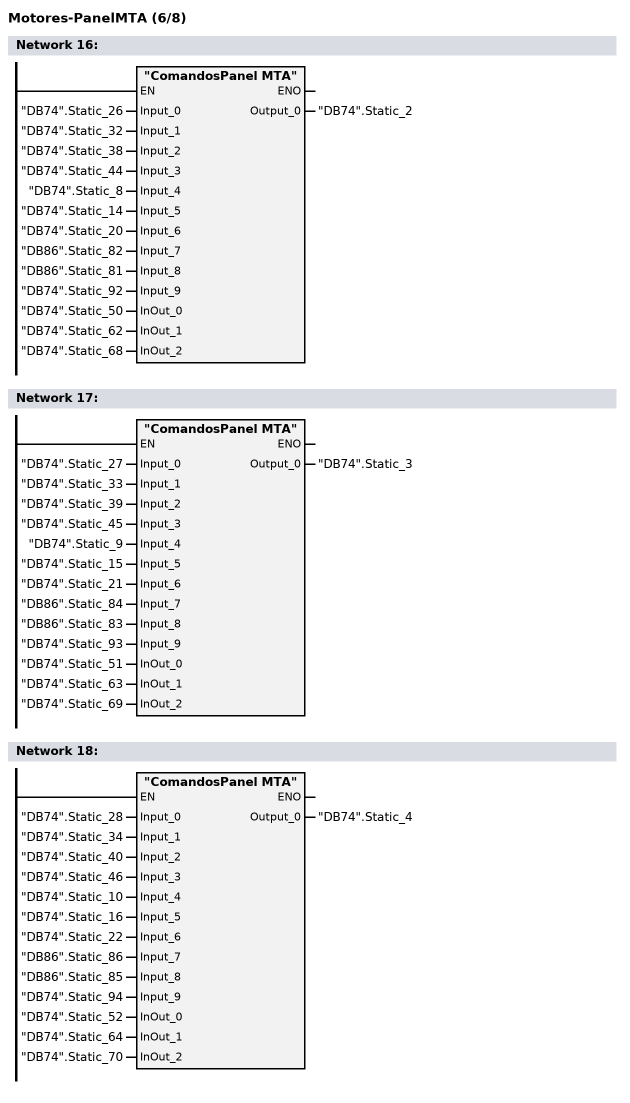
   RUNG wire#powerrail
      "ComandosPanel MTA"(Input_0 := "DB74".Static_26, Input_1 := "DB74".Static_32, Input_2 := "DB74".Static_38, Input_3 := "DB74".Static_44, Input_4 := "DB74".Static_8, Input_5 := "DB74".Static_14, Input_6 := "DB74".Static_20, Input_7 := "DB86".Static_82, Input_8 := "DB86".Static_81, Input_9 := "DB74".Static_92, Output_0 => "DB74".Static_2, InOut_0 := "DB74".Static_50, InOut_1 := "DB74".Static_62, InOut_2 := "DB74".Static_68)
   END_RUNG
   // the same network as SCL:
   "ComandosPanel MTA"(Input_0 := "DB74".Static_26,
                       Input_1 := "DB74".Static_32,
                       Input_2 := "DB74".Static_38,
                       Input_3 := "DB74".Static_44,
                       Input_4 := "DB74".Static_8,
                       Input_5 := "DB74".Static_14,
                       Input_6 := "DB74".Static_20,
                       Input_7 := "DB86".Static_82,
                       Input_8 := "DB86".Static_81,
                       Input_9 := "DB74".Static_92,
                       InOut_0 := "DB74".Static_50,
                       InOut_1 := "DB74".Static_62,
                       InOut_2 := "DB74".Static_68,
                       Output_0 => "DB74".Static_2);
END_REGION

REGION Network 17
   RUNG wire#powerrail
      "ComandosPanel MTA"(Input_0 := "DB74".Static_27, Input_1 := "DB74".Static_33, Input_2 := "DB74".Static_39, Input_3 := "DB74".Static_45, Input_4 := "DB74".Static_9, Input_5 := "DB74".Static_15, Input_6 := "DB74".Static_21, Input_7 := "DB86".Static_84, Input_8 := "DB86".Static_83, Input_9 := "DB74".Static_93, Output_0 => "DB74".Static_3, InOut_0 := "DB74".Static_51, InOut_1 := "DB74".Static_63, InOut_2 := "DB74".Static_69)
   END_RUNG
   // the same network as SCL:
   "ComandosPanel MTA"(Input_0 := "DB74".Static_27,
                       Input_1 := "DB74".Static_33,
                       Input_2 := "DB74".Static_39,
                       Input_3 := "DB74".Static_45,
                       Input_4 := "DB74".Static_9,
                       Input_5 := "DB74".Static_15,
                       Input_6 := "DB74".Static_21,
                       Input_7 := "DB86".Static_84,
                       Input_8 := "DB86".Static_83,
                       Input_9 := "DB74".Static_93,
                       InOut_0 := "DB74".Static_51,
                       InOut_1 := "DB74".Static_63,
                       InOut_2 := "DB74".Static_69,
                       Output_0 => "DB74".Static_3);
END_REGION

REGION Network 18
   RUNG wire#powerrail
      "ComandosPanel MTA"(Input_0 := "DB74".Static_28, Input_1 := "DB74".Static_34, Input_2 := "DB74".Static_40, Input_3 := "DB74".Static_46, Input_4 := "DB74".Static_10, Input_5 := "DB74".Static_16, Input_6 := "DB74".Static_22, Input_7 := "DB86".Static_86, Input_8 := "DB86".Static_85, Input_9 := "DB74".Static_94, Output_0 => "DB74".Static_4, InOut_0 := "DB74".Static_52, InOut_1 := "DB74".Static_64, InOut_2 := "DB74".Static_70)
   END_RUNG
   // the same network as SCL:
   "ComandosPanel MTA"(Input_0 := "DB74".Static_28,
                       Input_1 := "DB74".Static_34,
                       Input_2 := "DB74".Static_40,
                       Input_3 := "DB74".Static_46,
                       Input_4 := "DB74".Static_10,
                       Input_5 := "DB74".Static_16,
                       Input_6 := "DB74".Static_22,
                       Input_7 := "DB86".Static_86,
                       Input_8 := "DB86".Static_85,
                       Input_9 := "DB74".Static_94,
                       InOut_0 := "DB74".Static_52,
                       InOut_1 := "DB74".Static_64,
                       InOut_2 := "DB74".Static_70,
                       Output_0 => "DB74".Static_4);
END_REGION

REGION Network 19
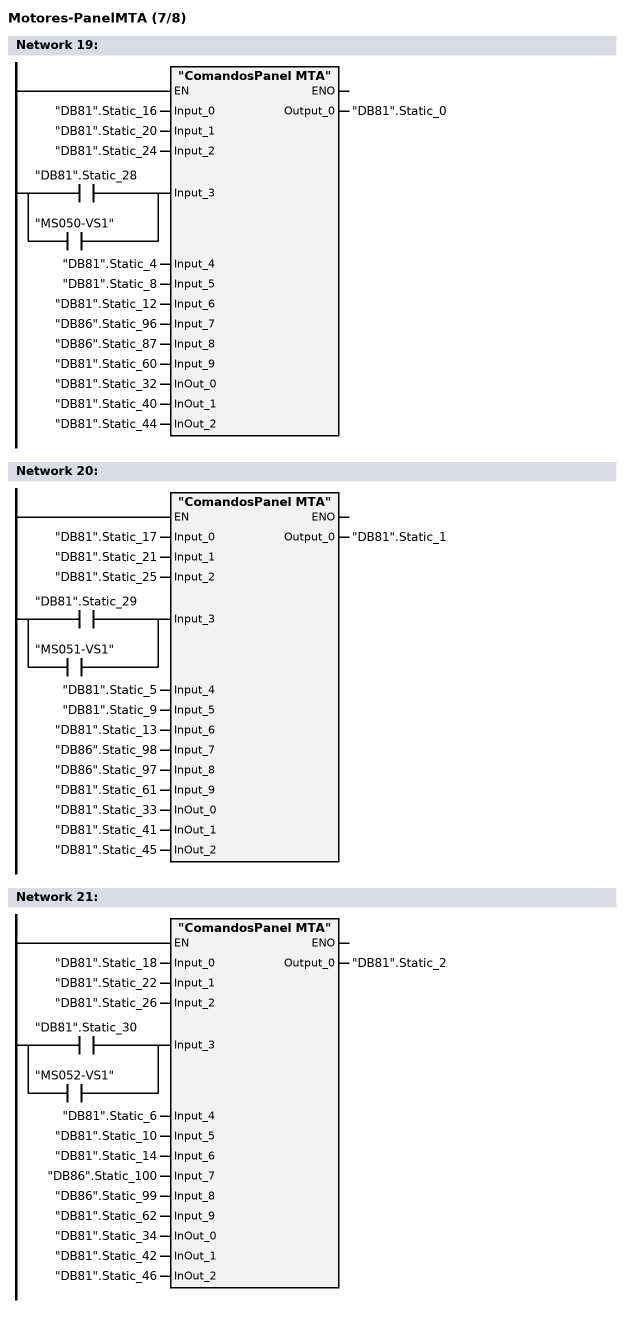
   RUNG wire#powerrail
      "ComandosPanel MTA"(Input_0 := "DB81".Static_16, Input_1 := "DB81".Static_20, Input_2 := "DB81".Static_24, Input_3 := wire#w1, Input_4 := "DB81".Static_4, Input_5 := "DB81".Static_8, Input_6 := "DB81".Static_12, Input_7 := "DB86".Static_96, Input_8 := "DB86".Static_87, Input_9 := "DB81".Static_60, Output_0 => "DB81".Static_0, InOut_0 := "DB81".Static_32, InOut_1 := "DB81".Static_40, InOut_2 := "DB81".Static_44)
   END_RUNG
   RUNG wire#powerrail
      Contact( "DB81".Static_28 )
   END_RUNG wire#w1
   RUNG wire#powerrail
      Contact( "MS050-VS1" )
   END_RUNG wire#w1
   // the same network as SCL:
   "ComandosPanel MTA"(Input_0 := "DB81".Static_16,
                       Input_1 := "DB81".Static_20,
                       Input_2 := "DB81".Static_24,
                       Input_3 := "DB81".Static_28 OR "MS050-VS1",
                       Input_4 := "DB81".Static_4,
                       Input_5 := "DB81".Static_8,
                       Input_6 := "DB81".Static_12,
                       Input_7 := "DB86".Static_96,
                       Input_8 := "DB86".Static_87,
                       Input_9 := "DB81".Static_60,
                       InOut_0 := "DB81".Static_32,
                       InOut_1 := "DB81".Static_40,
                       InOut_2 := "DB81".Static_44,
                       Output_0 => "DB81".Static_0);
END_REGION

REGION Network 20
   RUNG wire#powerrail
      "ComandosPanel MTA"(Input_0 := "DB81".Static_17, Input_1 := "DB81".Static_21, Input_2 := "DB81".Static_25, Input_3 := wire#w1, Input_4 := "DB81".Static_5, Input_5 := "DB81".Static_9, Input_6 := "DB81".Static_13, Input_7 := "DB86".Static_98, Input_8 := "DB86".Static_97, Input_9 := "DB81".Static_61, Output_0 => "DB81".Static_1, InOut_0 := "DB81".Static_33, InOut_1 := "DB81".Static_41, InOut_2 := "DB81".Static_45)
   END_RUNG
   RUNG wire#powerrail
      Contact( "DB81".Static_29 )
   END_RUNG wire#w1
   RUNG wire#powerrail
      Contact( "MS051-VS1" )
   END_RUNG wire#w1
   // the same network as SCL:
   "ComandosPanel MTA"(Input_0 := "DB81".Static_17,
                       Input_1 := "DB81".Static_21,
                       Input_2 := "DB81".Static_25,
                       Input_3 := "DB81".Static_29 OR "MS051-VS1",
                       Input_4 := "DB81".Static_5,
                       Input_5 := "DB81".Static_9,
                       Input_6 := "DB81".Static_13,
                       Input_7 := "DB86".Static_98,
                       Input_8 := "DB86".Static_97,
                       Input_9 := "DB81".Static_61,
                       InOut_0 := "DB81".Static_33,
                       InOut_1 := "DB81".Static_41,
                       InOut_2 := "DB81".Static_45,
                       Output_0 => "DB81".Static_1);
END_REGION

REGION Network 21
   RUNG wire#powerrail
      "ComandosPanel MTA"(Input_0 := "DB81".Static_18, Input_1 := "DB81".Static_22, Input_2 := "DB81".Static_26, Input_3 := wire#w1, Input_4 := "DB81".Static_6, Input_5 := "DB81".Static_10, Input_6 := "DB81".Static_14, Input_7 := "DB86".Static_100, Input_8 := "DB86".Static_99, Input_9 := "DB81".Static_62, Output_0 => "DB81".Static_2, InOut_0 := "DB81".Static_34, InOut_1 := "DB81".Static_42, InOut_2 := "DB81".Static_46)
   END_RUNG
   RUNG wire#powerrail
      Contact( "DB81".Static_30 )
   END_RUNG wire#w1
   RUNG wire#powerrail
      Contact( "MS052-VS1" )
   END_RUNG wire#w1
   // the same network as SCL:
   "ComandosPanel MTA"(Input_0 := "DB81".Static_18,
                       Input_1 := "DB81".Static_22,
                       Input_2 := "DB81".Static_26,
                       Input_3 := "DB81".Static_30 OR "MS052-VS1",
                       Input_4 := "DB81".Static_6,
                       Input_5 := "DB81".Static_10,
                       Input_6 := "DB81".Static_14,
                       Input_7 := "DB86".Static_100,
                       Input_8 := "DB86".Static_99,
                       Input_9 := "DB81".Static_62,
                       InOut_0 := "DB81".Static_34,
                       InOut_1 := "DB81".Static_42,
                       InOut_2 := "DB81".Static_46,
                       Output_0 => "DB81".Static_2);
END_REGION

REGION Network 22
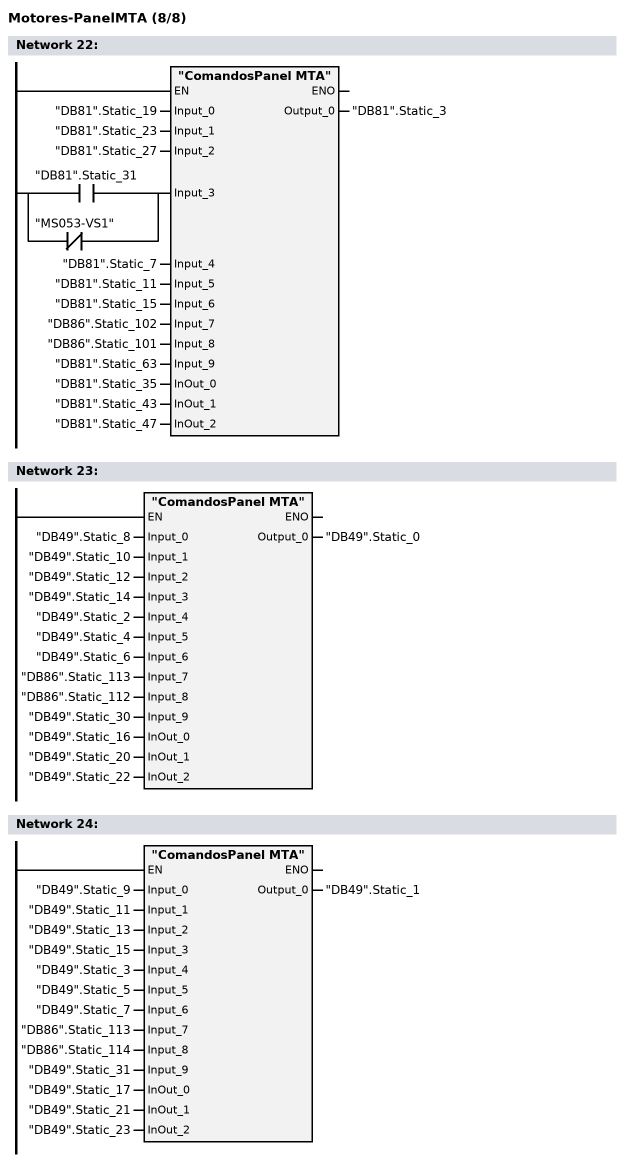
   RUNG wire#powerrail
      "ComandosPanel MTA"(Input_0 := "DB81".Static_19, Input_1 := "DB81".Static_23, Input_2 := "DB81".Static_27, Input_3 := wire#w1, Input_4 := "DB81".Static_7, Input_5 := "DB81".Static_11, Input_6 := "DB81".Static_15, Input_7 := "DB86".Static_102, Input_8 := "DB86".Static_101, Input_9 := "DB81".Static_63, Output_0 => "DB81".Static_3, InOut_0 := "DB81".Static_35, InOut_1 := "DB81".Static_43, InOut_2 := "DB81".Static_47)
   END_RUNG
   RUNG wire#powerrail
      Contact( "DB81".Static_31 )
   END_RUNG wire#w1
   RUNG wire#powerrail
      I_Contact( "MS053-VS1" )
   END_RUNG wire#w1
   // the same network as SCL:
   "ComandosPanel MTA"(Input_0 := "DB81".Static_19,
                       Input_1 := "DB81".Static_23,
                       Input_2 := "DB81".Static_27,
                       Input_3 := "DB81".Static_31 OR NOT "MS053-VS1",
                       Input_4 := "DB81".Static_7,
                       Input_5 := "DB81".Static_11,
                       Input_6 := "DB81".Static_15,
                       Input_7 := "DB86".Static_102,
                       Input_8 := "DB86".Static_101,
                       Input_9 := "DB81".Static_63,
                       InOut_0 := "DB81".Static_35,
                       InOut_1 := "DB81".Static_43,
                       InOut_2 := "DB81".Static_47,
                       Output_0 => "DB81".Static_3);
END_REGION

REGION Network 23
   RUNG wire#powerrail
      "ComandosPanel MTA"(Input_0 := "DB49".Static_8, Input_1 := "DB49".Static_10, Input_2 := "DB49".Static_12, Input_3 := "DB49".Static_14, Input_4 := "DB49".Static_2, Input_5 := "DB49".Static_4, Input_6 := "DB49".Static_6, Input_7 := "DB86".Static_113, Input_8 := "DB86".Static_112, Input_9 := "DB49".Static_30, Output_0 => "DB49".Static_0, InOut_0 := "DB49".Static_16, InOut_1 := "DB49".Static_20, InOut_2 := "DB49".Static_22)
   END_RUNG
   // the same network as SCL:
   "ComandosPanel MTA"(Input_0 := "DB49".Static_8,
                       Input_1 := "DB49".Static_10,
                       Input_2 := "DB49".Static_12,
                       Input_3 := "DB49".Static_14,
                       Input_4 := "DB49".Static_2,
                       Input_5 := "DB49".Static_4,
                       Input_6 := "DB49".Static_6,
                       Input_7 := "DB86".Static_113,
                       Input_8 := "DB86".Static_112,
                       Input_9 := "DB49".Static_30,
                       InOut_0 := "DB49".Static_16,
                       InOut_1 := "DB49".Static_20,
                       InOut_2 := "DB49".Static_22,
                       Output_0 => "DB49".Static_0);
END_REGION

REGION Network 24
   RUNG wire#powerrail
      "ComandosPanel MTA"(Input_0 := "DB49".Static_9, Input_1 := "DB49".Static_11, Input_2 := "DB49".Static_13, Input_3 := "DB49".Static_15, Input_4 := "DB49".Static_3, Input_5 := "DB49".Static_5, Input_6 := "DB49".Static_7, Input_7 := "DB86".Static_113, Input_8 := "DB86".Static_114, Input_9 := "DB49".Static_31, Output_0 => "DB49".Static_1, InOut_0 := "DB49".Static_17, InOut_1 := "DB49".Static_21, InOut_2 := "DB49".Static_23)
   END_RUNG
   // the same network as SCL:
   "ComandosPanel MTA"(Input_0 := "DB49".Static_9,
                       Input_1 := "DB49".Static_11,
                       Input_2 := "DB49".Static_13,
                       Input_3 := "DB49".Static_15,
                       Input_4 := "DB49".Static_3,
                       Input_5 := "DB49".Static_5,
                       Input_6 := "DB49".Static_7,
                       Input_7 := "DB86".Static_113,
                       Input_8 := "DB86".Static_114,
                       Input_9 := "DB49".Static_31,
                       InOut_0 := "DB49".Static_17,
                       InOut_1 := "DB49".Static_21,
                       InOut_2 := "DB49".Static_23,
                       Output_0 => "DB49".Static_1);
END_REGION
END_FUNCTION

FUNCTION "ComandosPanel MTA" : Void   // FC19, LAD
{ S7_Optimized_Access := 'FALSE' }
VERSION : 0.1
   VAR_TEMP   // added for the SCL form of the ladder/FBD networks
      _w1 : Bool;
   END_VAR
BEGIN

REGION Network 1
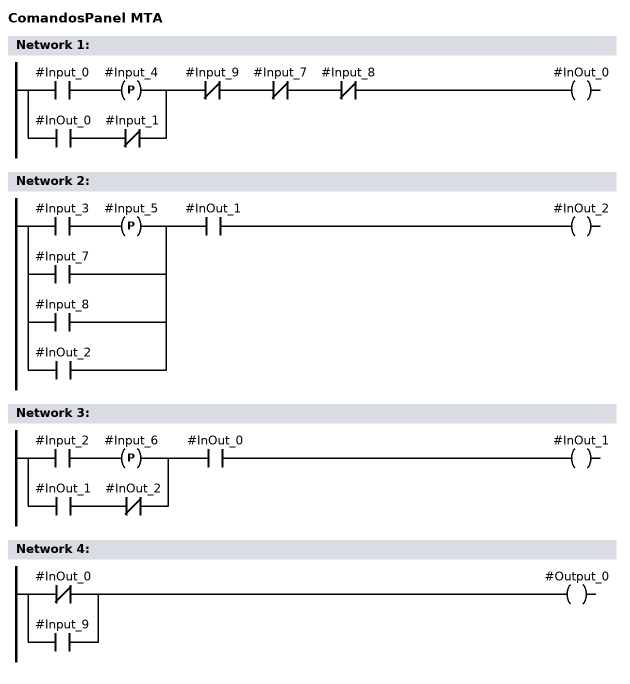
   RUNG wire#powerrail
      Contact( #Input_0 )
      P_Trig( #Input_4 )
      wire#w1
      I_Contact( #Input_9 )
      I_Contact( #Input_7 )
      I_Contact( #Input_8 )
      Coil( #InOut_0 )
   END_RUNG
   RUNG wire#powerrail
      Contact( #InOut_0 )
      I_Contact( #Input_1 )
   END_RUNG wire#w1
   // the same network as SCL:
   #_w1 := #Input_0 AND NOT #Input_4;   // rising edge
   #Input_4 := #Input_0;
   #InOut_0 := (#_w1 OR (#InOut_0 AND NOT #Input_1)) AND NOT #Input_9 AND NOT #Input_7 AND NOT #Input_8;
END_REGION

REGION Network 2
   RUNG wire#powerrail
      Contact( #Input_3 )
      P_Trig( #Input_5 )
      wire#w1
      Contact( #InOut_1 )
      Coil( #InOut_2 )
   END_RUNG
   RUNG wire#powerrail
      Contact( #Input_7 )
   END_RUNG wire#w1
   RUNG wire#powerrail
      Contact( #Input_8 )
   END_RUNG wire#w1
   RUNG wire#powerrail
      Contact( #InOut_2 )
   END_RUNG wire#w1
   // the same network as SCL:
   #_w1 := #Input_3 AND NOT #Input_5;   // rising edge
   #Input_5 := #Input_3;
   #InOut_2 := (#_w1 OR #Input_7 OR #Input_8 OR #InOut_2) AND #InOut_1;
END_REGION

REGION Network 3
   RUNG wire#powerrail
      Contact( #Input_2 )
      P_Trig( #Input_6 )
      wire#w1
      Contact( #InOut_0 )
      Coil( #InOut_1 )
   END_RUNG
   RUNG wire#powerrail
      Contact( #InOut_1 )
      I_Contact( #InOut_2 )
   END_RUNG wire#w1
   // the same network as SCL:
   #_w1 := #Input_2 AND NOT #Input_6;   // rising edge
   #Input_6 := #Input_2;
   #InOut_1 := (#_w1 OR (#InOut_1 AND NOT #InOut_2)) AND #InOut_0;
END_REGION

REGION Network 4
   RUNG wire#powerrail
      I_Contact( #InOut_0 )
      wire#w1
      Coil( #Output_0 )
   END_RUNG
   RUNG wire#powerrail
      Contact( #Input_9 )
   END_RUNG wire#w1
   // the same network as SCL:
   #Output_0 := NOT #InOut_0 OR #Input_9;
END_REGION
END_FUNCTION

FUNCTION "FC-ANIM-CMP" : Void   // FC43, LAD
{ S7_Optimized_Access := 'FALSE' }
VERSION : 0.1
BEGIN

REGION Network 1
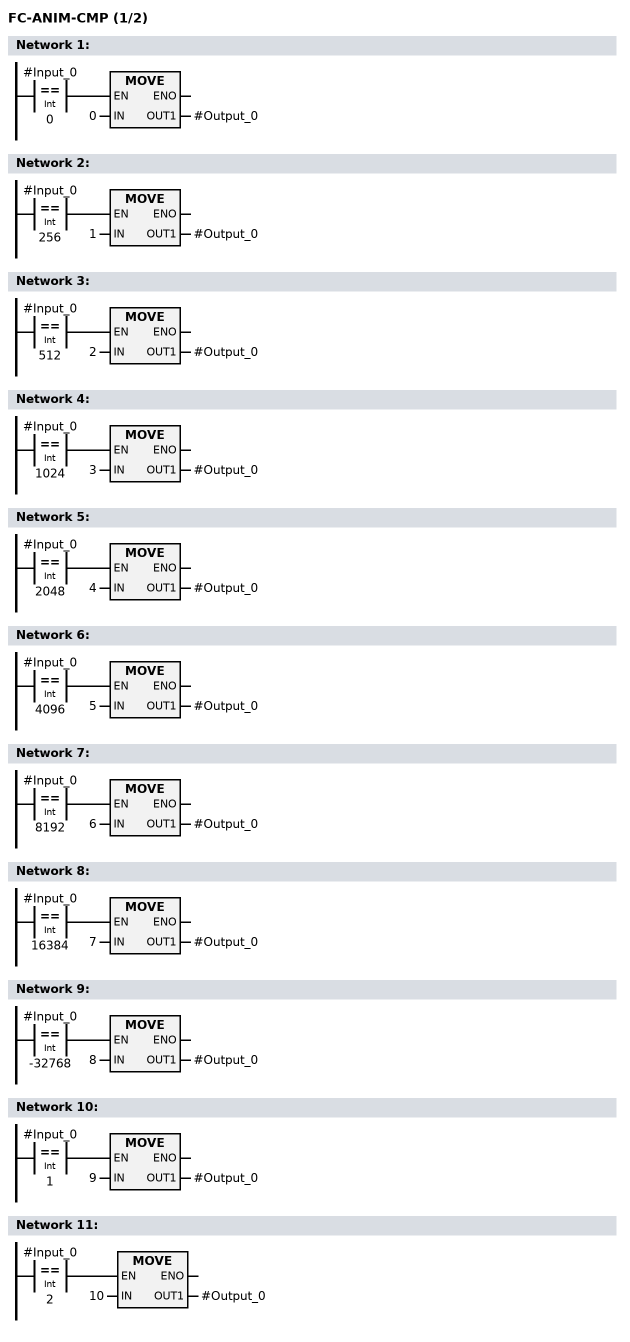
   RUNG wire#powerrail
      { S7_Templates := "SrcType := Int" } EQ_Contact(in1 := #Input_0, in2 := 0)
      { S7_GenerateENO := "TRUE" } Move(in := 0, out1 => #Output_0)
   END_RUNG
   // the same network as SCL:
   IF #Input_0 = 0 THEN #Output_0 := 0; END_IF;
END_REGION

REGION Network 2
   RUNG wire#powerrail
      { S7_Templates := "SrcType := Int" } EQ_Contact(in1 := #Input_0, in2 := 256)
      { S7_GenerateENO := "TRUE" } Move(in := 1, out1 => #Output_0)
   END_RUNG
   // the same network as SCL:
   IF #Input_0 = 256 THEN #Output_0 := 1; END_IF;
END_REGION

REGION Network 3
   RUNG wire#powerrail
      { S7_Templates := "SrcType := Int" } EQ_Contact(in1 := #Input_0, in2 := 512)
      { S7_GenerateENO := "TRUE" } Move(in := 2, out1 => #Output_0)
   END_RUNG
   // the same network as SCL:
   IF #Input_0 = 512 THEN #Output_0 := 2; END_IF;
END_REGION

REGION Network 4
   RUNG wire#powerrail
      { S7_Templates := "SrcType := Int" } EQ_Contact(in1 := #Input_0, in2 := 1024)
      { S7_GenerateENO := "TRUE" } Move(in := 3, out1 => #Output_0)
   END_RUNG
   // the same network as SCL:
   IF #Input_0 = 1024 THEN #Output_0 := 3; END_IF;
END_REGION

REGION Network 5
   RUNG wire#powerrail
      { S7_Templates := "SrcType := Int" } EQ_Contact(in1 := #Input_0, in2 := 2048)
      { S7_GenerateENO := "TRUE" } Move(in := 4, out1 => #Output_0)
   END_RUNG
   // the same network as SCL:
   IF #Input_0 = 2048 THEN #Output_0 := 4; END_IF;
END_REGION

REGION Network 6
   RUNG wire#powerrail
      { S7_Templates := "SrcType := Int" } EQ_Contact(in1 := #Input_0, in2 := 4096)
      { S7_GenerateENO := "TRUE" } Move(in := 5, out1 => #Output_0)
   END_RUNG
   // the same network as SCL:
   IF #Input_0 = 4096 THEN #Output_0 := 5; END_IF;
END_REGION

REGION Network 7
   RUNG wire#powerrail
      { S7_Templates := "SrcType := Int" } EQ_Contact(in1 := #Input_0, in2 := 8192)
      { S7_GenerateENO := "TRUE" } Move(in := 6, out1 => #Output_0)
   END_RUNG
   // the same network as SCL:
   IF #Input_0 = 8192 THEN #Output_0 := 6; END_IF;
END_REGION

REGION Network 8
   RUNG wire#powerrail
      { S7_Templates := "SrcType := Int" } EQ_Contact(in1 := #Input_0, in2 := 16384)
      { S7_GenerateENO := "TRUE" } Move(in := 7, out1 => #Output_0)
   END_RUNG
   // the same network as SCL:
   IF #Input_0 = 16384 THEN #Output_0 := 7; END_IF;
END_REGION

REGION Network 9
   RUNG wire#powerrail
      { S7_Templates := "SrcType := Int" } EQ_Contact(in1 := #Input_0, in2 := -32768)
      { S7_GenerateENO := "TRUE" } Move(in := 8, out1 => #Output_0)
   END_RUNG
   // the same network as SCL:
   IF #Input_0 = (-32768) THEN #Output_0 := 8; END_IF;
END_REGION

REGION Network 10
   RUNG wire#powerrail
      { S7_Templates := "SrcType := Int" } EQ_Contact(in1 := #Input_0, in2 := 1)
      { S7_GenerateENO := "TRUE" } Move(in := 9, out1 => #Output_0)
   END_RUNG
   // the same network as SCL:
   IF #Input_0 = 1 THEN #Output_0 := 9; END_IF;
END_REGION

REGION Network 11
   RUNG wire#powerrail
      { S7_Templates := "SrcType := Int" } EQ_Contact(in1 := #Input_0, in2 := 2)
      { S7_GenerateENO := "TRUE" } Move(in := 10, out1 => #Output_0)
   END_RUNG
   // the same network as SCL:
   IF #Input_0 = 2 THEN #Output_0 := 10; END_IF;
END_REGION

REGION Network 12
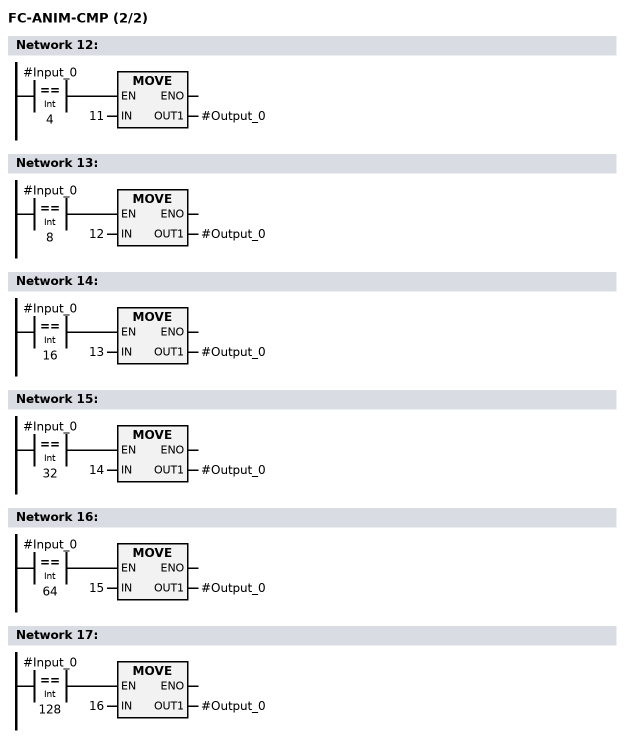
   RUNG wire#powerrail
      { S7_Templates := "SrcType := Int" } EQ_Contact(in1 := #Input_0, in2 := 4)
      { S7_GenerateENO := "TRUE" } Move(in := 11, out1 => #Output_0)
   END_RUNG
   // the same network as SCL:
   IF #Input_0 = 4 THEN #Output_0 := 11; END_IF;
END_REGION

REGION Network 13
   RUNG wire#powerrail
      { S7_Templates := "SrcType := Int" } EQ_Contact(in1 := #Input_0, in2 := 8)
      { S7_GenerateENO := "TRUE" } Move(in := 12, out1 => #Output_0)
   END_RUNG
   // the same network as SCL:
   IF #Input_0 = 8 THEN #Output_0 := 12; END_IF;
END_REGION

REGION Network 14
   RUNG wire#powerrail
      { S7_Templates := "SrcType := Int" } EQ_Contact(in1 := #Input_0, in2 := 16)
      { S7_GenerateENO := "TRUE" } Move(in := 13, out1 => #Output_0)
   END_RUNG
   // the same network as SCL:
   IF #Input_0 = 16 THEN #Output_0 := 13; END_IF;
END_REGION

REGION Network 15
   RUNG wire#powerrail
      { S7_Templates := "SrcType := Int" } EQ_Contact(in1 := #Input_0, in2 := 32)
      { S7_GenerateENO := "TRUE" } Move(in := 14, out1 => #Output_0)
   END_RUNG
   // the same network as SCL:
   IF #Input_0 = 32 THEN #Output_0 := 14; END_IF;
END_REGION

REGION Network 16
   RUNG wire#powerrail
      { S7_Templates := "SrcType := Int" } EQ_Contact(in1 := #Input_0, in2 := 64)
      { S7_GenerateENO := "TRUE" } Move(in := 15, out1 => #Output_0)
   END_RUNG
   // the same network as SCL:
   IF #Input_0 = 64 THEN #Output_0 := 15; END_IF;
END_REGION

REGION Network 17
   RUNG wire#powerrail
      { S7_Templates := "SrcType := Int" } EQ_Contact(in1 := #Input_0, in2 := 128)
      { S7_GenerateENO := "TRUE" } Move(in := 16, out1 => #Output_0)
   END_RUNG
   // the same network as SCL:
   IF #Input_0 = 128 THEN #Output_0 := 16; END_IF;
END_REGION
END_FUNCTION

// folder: Secadoras/Alta

FUNCTION "EnclavSecAltaMTA" : Void   // FC12, LAD
{ S7_Optimized_Access := 'FALSE' }
VERSION : 0.1
BEGIN

REGION Network 1
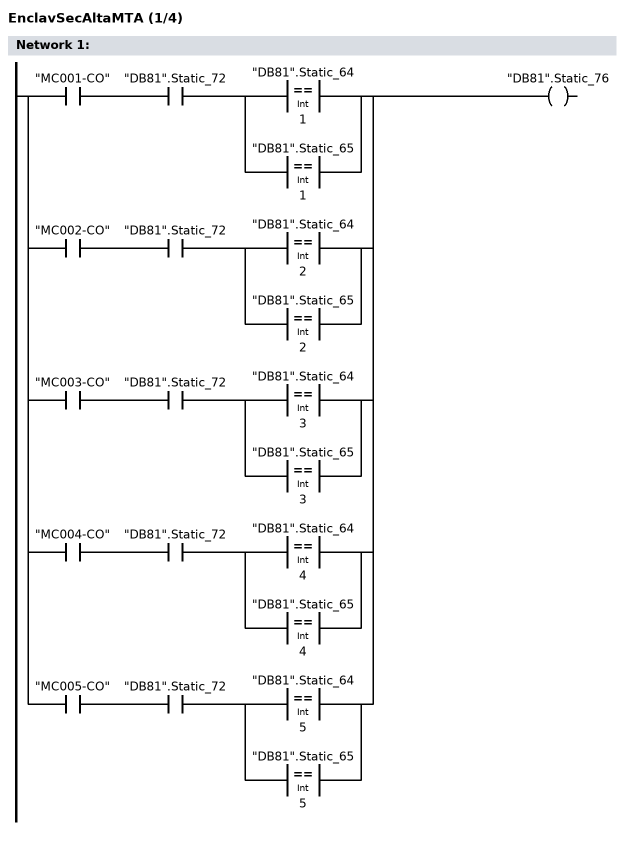
   "DB81".Static_76 := ("MC001-CO" AND "DB81".Static_72 AND (("DB81".Static_64 = 1) OR ("DB81".Static_65 = 1))) OR ("MC002-CO" AND "DB81".Static_72 AND (("DB81".Static_64 = 2) OR ("DB81".Static_65 = 2))) OR ("MC003-CO" AND "DB81".Static_72 AND (("DB81".Static_64 = 3) OR ("DB81".Static_65 = 3))) OR ("MC004-CO" AND "DB81".Static_72 AND (("DB81".Static_64 = 4) OR ("DB81".Static_65 = 4))) OR ("MC005-CO" AND "DB81".Static_72 AND (("DB81".Static_64 = 5) OR ("DB81".Static_65 = 5)));
END_REGION

REGION Network 2
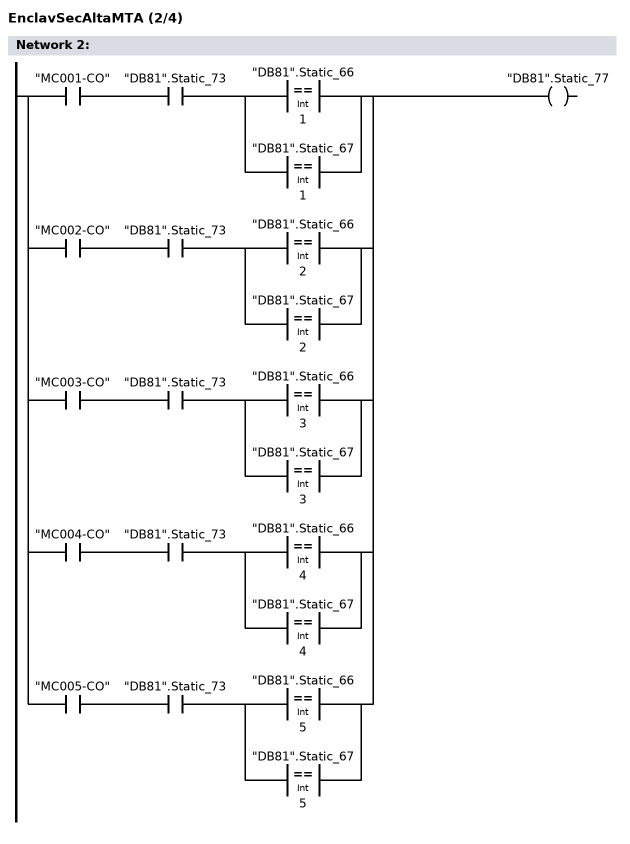
   "DB81".Static_77 := ("MC001-CO" AND "DB81".Static_73 AND (("DB81".Static_66 = 1) OR ("DB81".Static_67 = 1))) OR ("MC002-CO" AND "DB81".Static_73 AND (("DB81".Static_66 = 2) OR ("DB81".Static_67 = 2))) OR ("MC003-CO" AND "DB81".Static_73 AND (("DB81".Static_66 = 3) OR ("DB81".Static_67 = 3))) OR ("MC004-CO" AND "DB81".Static_73 AND (("DB81".Static_66 = 4) OR ("DB81".Static_67 = 4))) OR ("MC005-CO" AND "DB81".Static_73 AND (("DB81".Static_66 = 5) OR ("DB81".Static_67 = 5)));
END_REGION

REGION Network 3
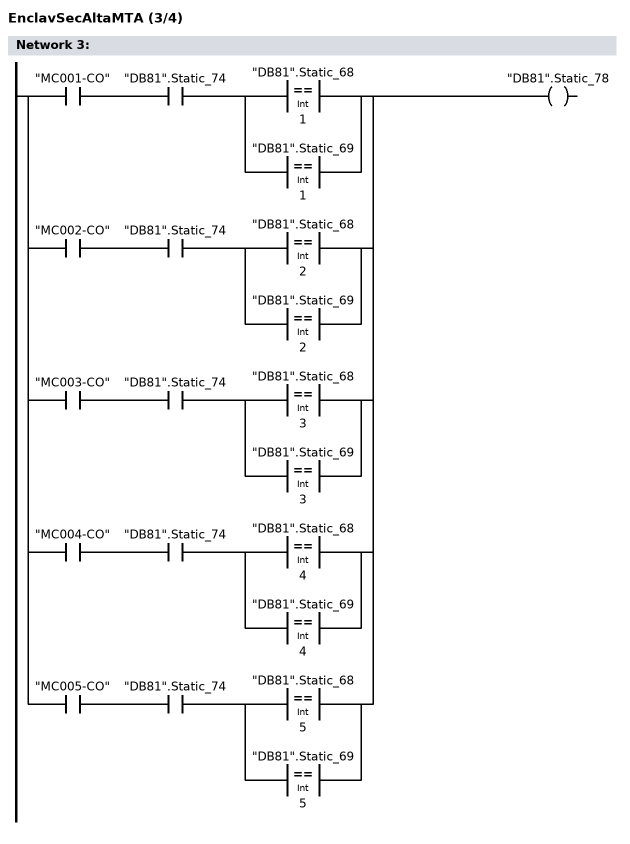
   "DB81".Static_78 := ("MC001-CO" AND "DB81".Static_74 AND (("DB81".Static_68 = 1) OR ("DB81".Static_69 = 1))) OR ("MC002-CO" AND "DB81".Static_74 AND (("DB81".Static_68 = 2) OR ("DB81".Static_69 = 2))) OR ("MC003-CO" AND "DB81".Static_74 AND (("DB81".Static_68 = 3) OR ("DB81".Static_69 = 3))) OR ("MC004-CO" AND "DB81".Static_74 AND (("DB81".Static_68 = 4) OR ("DB81".Static_69 = 4))) OR ("MC005-CO" AND "DB81".Static_74 AND (("DB81".Static_68 = 5) OR ("DB81".Static_69 = 5)));
END_REGION

REGION Network 4
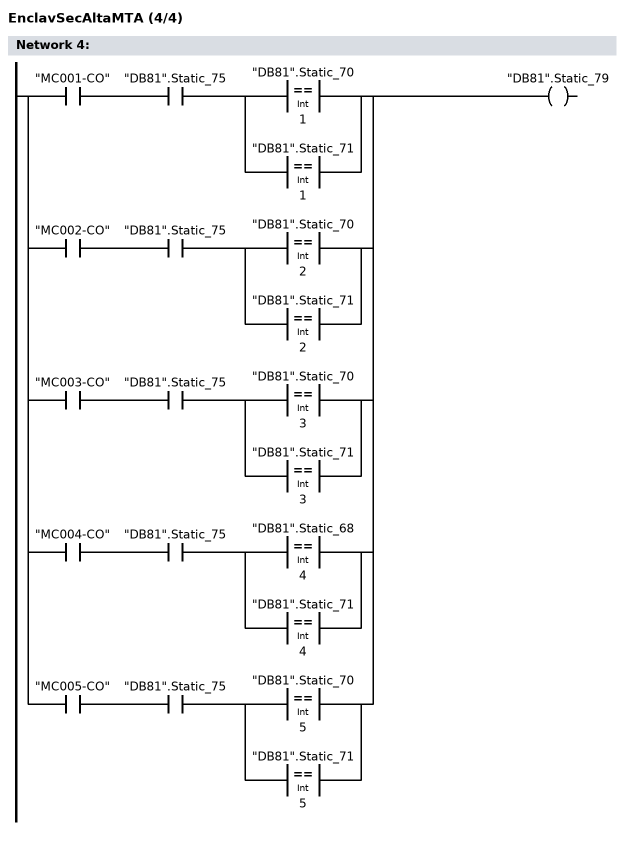
   "DB81".Static_79 := ("MC001-CO" AND "DB81".Static_75 AND (("DB81".Static_70 = 1) OR ("DB81".Static_71 = 1))) OR ("MC002-CO" AND "DB81".Static_75 AND (("DB81".Static_70 = 2) OR ("DB81".Static_71 = 2))) OR ("MC003-CO" AND "DB81".Static_75 AND (("DB81".Static_70 = 3) OR ("DB81".Static_71 = 3))) OR ("MC004-CO" AND "DB81".Static_75 AND (("DB81".Static_68 = 4) OR ("DB81".Static_71 = 4))) OR ("MC005-CO" AND "DB81".Static_75 AND (("DB81".Static_70 = 5) OR ("DB81".Static_71 = 5)));
END_REGION
END_FUNCTION

// folder: Torres de Agua/Cavaleto

FUNCTION "TorresCavaletoMTA" : Void   // FC14, LAD
{ S7_Optimized_Access := 'FALSE' }
VERSION : 0.1
BEGIN

REGION Network 1
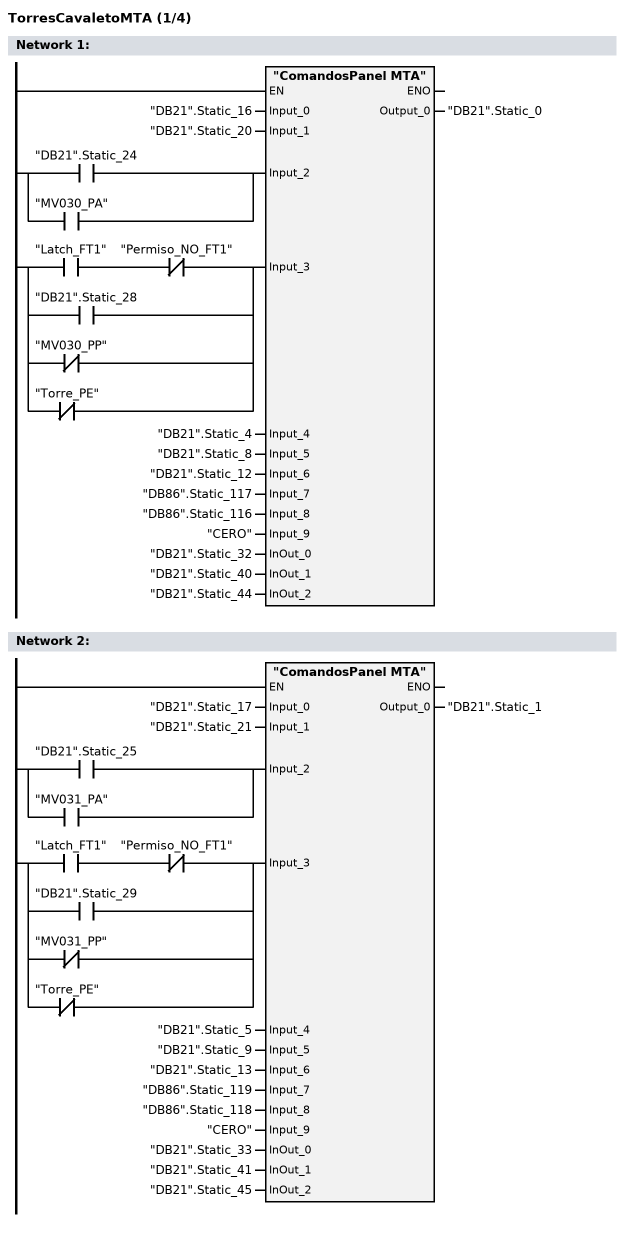
   "ComandosPanel MTA"(Input_0 := "DB21".Static_16,
                       Input_1 := "DB21".Static_20,
                       Input_2 := "DB21".Static_24 OR "MV030_PA",
                       Input_3 := "DB21".Static_28 OR NOT "MV030_PP" OR NOT "Torre_PE" OR ("Latch_FT1" AND NOT "Permiso_NO_FT1"),
                       Input_4 := "DB21".Static_4,
                       Input_5 := "DB21".Static_8,
                       Input_6 := "DB21".Static_12,
                       Input_7 := "DB86".Static_117,
                       Input_8 := "DB86".Static_116,
                       Input_9 := "CERO",
                       InOut_0 := "DB21".Static_32,
                       InOut_1 := "DB21".Static_40,
                       InOut_2 := "DB21".Static_44,
                       Output_0 => "DB21".Static_0);
END_REGION

REGION Network 2
   "ComandosPanel MTA"(Input_0 := "DB21".Static_17,
                       Input_1 := "DB21".Static_21,
                       Input_2 := "DB21".Static_25 OR "MV031_PA",
                       Input_3 := "DB21".Static_29 OR NOT "MV031_PP" OR NOT "Torre_PE" OR ("Latch_FT1" AND NOT "Permiso_NO_FT1"),
                       Input_4 := "DB21".Static_5,
                       Input_5 := "DB21".Static_9,
                       Input_6 := "DB21".Static_13,
                       Input_7 := "DB86".Static_119,
                       Input_8 := "DB86".Static_118,
                       Input_9 := "CERO",
                       InOut_0 := "DB21".Static_33,
                       InOut_1 := "DB21".Static_41,
                       InOut_2 := "DB21".Static_45,
                       Output_0 => "DB21".Static_1);
END_REGION

REGION Network 3
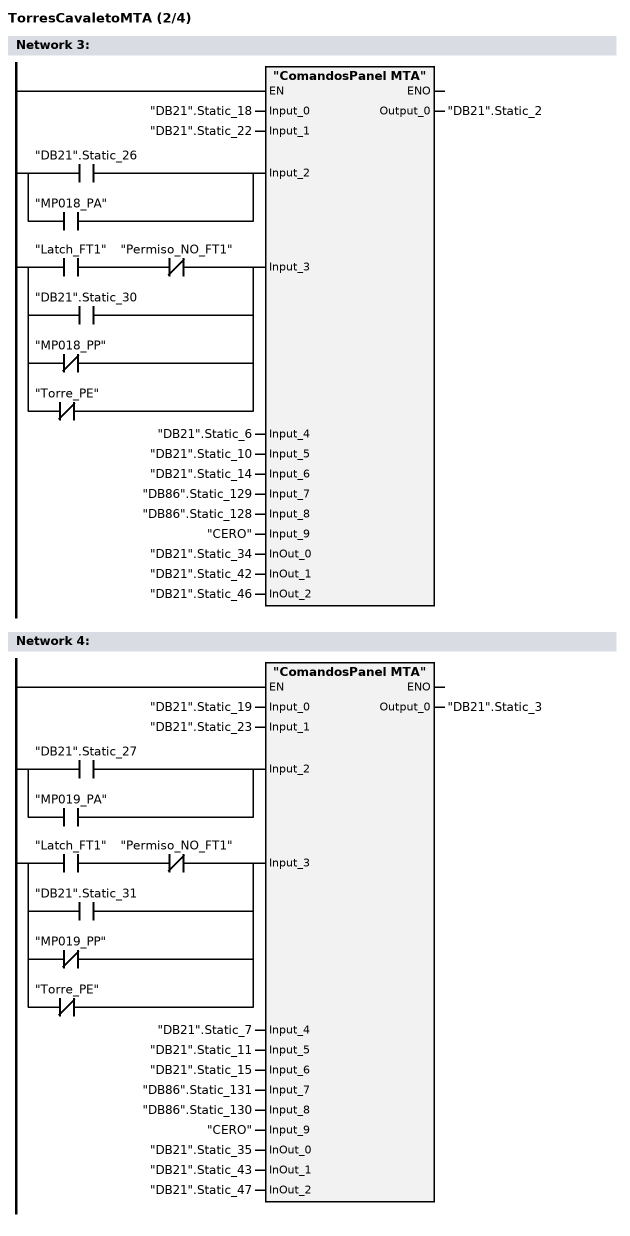
   "ComandosPanel MTA"(Input_0 := "DB21".Static_18,
                       Input_1 := "DB21".Static_22,
                       Input_2 := "DB21".Static_26 OR "MP018_PA",
                       Input_3 := "DB21".Static_30 OR NOT "MP018_PP" OR NOT "Torre_PE" OR ("Latch_FT1" AND NOT "Permiso_NO_FT1"),
                       Input_4 := "DB21".Static_6,
                       Input_5 := "DB21".Static_10,
                       Input_6 := "DB21".Static_14,
                       Input_7 := "DB86".Static_129,
                       Input_8 := "DB86".Static_128,
                       Input_9 := "CERO",
                       InOut_0 := "DB21".Static_34,
                       InOut_1 := "DB21".Static_42,
                       InOut_2 := "DB21".Static_46,
                       Output_0 => "DB21".Static_2);
END_REGION

REGION Network 4
   "ComandosPanel MTA"(Input_0 := "DB21".Static_19,
                       Input_1 := "DB21".Static_23,
                       Input_2 := "DB21".Static_27 OR "MP019_PA",
                       Input_3 := "DB21".Static_31 OR NOT "MP019_PP" OR NOT "Torre_PE" OR ("Latch_FT1" AND NOT "Permiso_NO_FT1"),
                       Input_4 := "DB21".Static_7,
                       Input_5 := "DB21".Static_11,
                       Input_6 := "DB21".Static_15,
                       Input_7 := "DB86".Static_131,
                       Input_8 := "DB86".Static_130,
                       Input_9 := "CERO",
                       InOut_0 := "DB21".Static_35,
                       InOut_1 := "DB21".Static_43,
                       InOut_2 := "DB21".Static_47,
                       Output_0 => "DB21".Static_3);
END_REGION

REGION Network 5
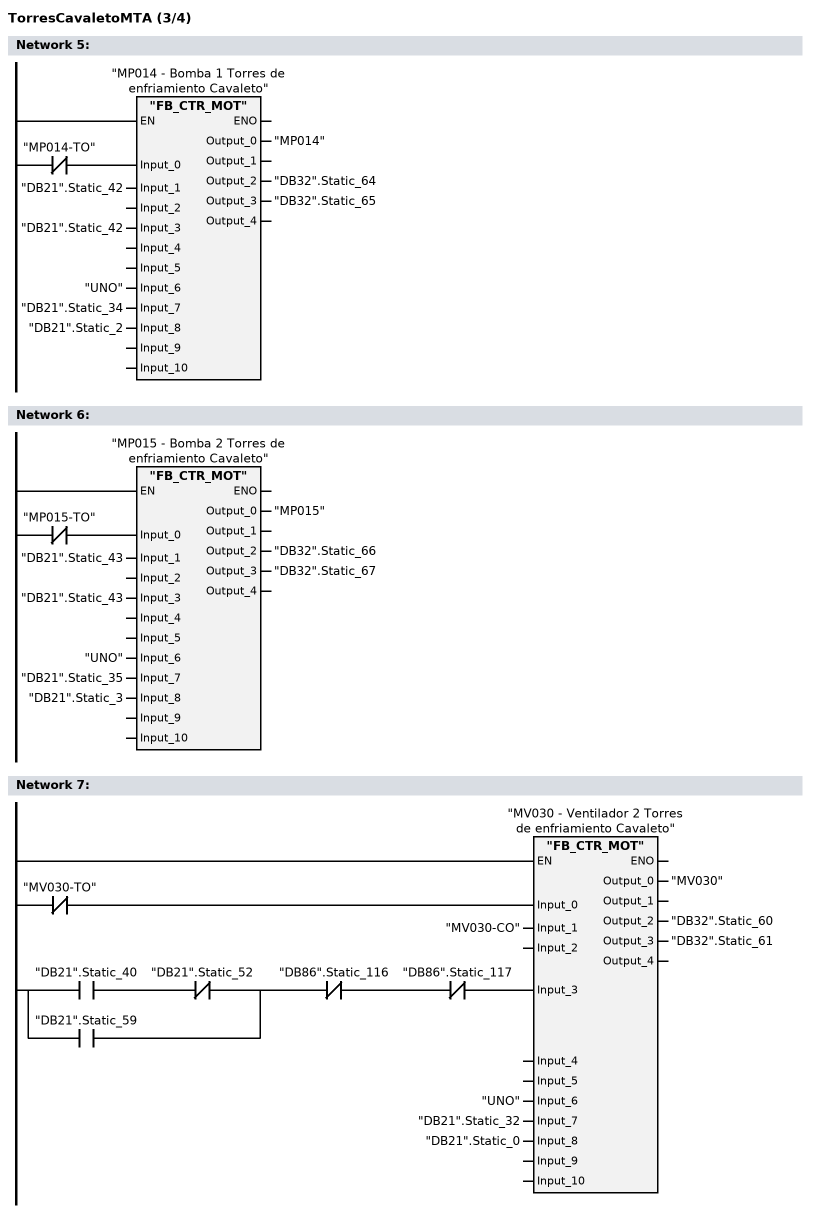
   RUNG wire#powerrail
      "MP014 - Bomba 1 Torres de enfriamiento Cavaleto"(Input_1 := "DB21".Static_42, Input_2 :=, Input_3 := "DB21".Static_42, Input_4 :=, Input_5 :=, Input_6 := "UNO", Input_7 := "DB21".Static_34, Input_8 := "DB21".Static_2, Input_9 :=, Input_10 :=, Output_0 => "MP014", Output_1 =>, Output_2 => "DB32".Static_64, Output_3 => "DB32".Static_65, Output_4 =>, Input_0 := wire#w1)
   END_RUNG
   RUNG wire#powerrail
      I_Contact( "MP014-TO" )
   END_RUNG wire#w1
   // the same network as SCL:
   "MP014 - Bomba 1 Torres de enfriamiento Cavaleto"(Input_0 := NOT "MP014-TO",   // "FB_CTR_MOT"
                           Input_1 := "DB21".Static_42,
                           Input_3 := "DB21".Static_42,
                           Input_6 := "UNO",
                           Input_7 := "DB21".Static_34,
                           Input_8 := "DB21".Static_2,
                           Output_0 => "MP014",
                           Output_2 => "DB32".Static_64,
                           Output_3 => "DB32".Static_65);
END_REGION

REGION Network 6
   RUNG wire#powerrail
      "MP015 - Bomba 2 Torres de enfriamiento Cavaleto"(Input_1 := "DB21".Static_43, Input_2 :=, Input_3 := "DB21".Static_43, Input_4 :=, Input_5 :=, Input_6 := "UNO", Input_7 := "DB21".Static_35, Input_8 := "DB21".Static_3, Input_9 :=, Input_10 :=, Output_0 => "MP015", Output_1 =>, Output_2 => "DB32".Static_66, Output_3 => "DB32".Static_67, Output_4 =>, Input_0 := wire#w1)
   END_RUNG
   RUNG wire#powerrail
      I_Contact( "MP015-TO" )
   END_RUNG wire#w1
   // the same network as SCL:
   "MP015 - Bomba 2 Torres de enfriamiento Cavaleto"(Input_0 := NOT "MP015-TO",   // "FB_CTR_MOT"
                           Input_1 := "DB21".Static_43,
                           Input_3 := "DB21".Static_43,
                           Input_6 := "UNO",
                           Input_7 := "DB21".Static_35,
                           Input_8 := "DB21".Static_3,
                           Output_0 => "MP015",
                           Output_2 => "DB32".Static_66,
                           Output_3 => "DB32".Static_67);
END_REGION

REGION Network 7
   "MV030 - Ventilador 2 Torres de enfriamiento Cavaleto"(Input_0 := NOT "MV030-TO",   // "FB_CTR_MOT"
                           Input_1 := "MV030-CO",
                           Input_3 := (("DB21".Static_40 AND NOT "DB21".Static_52) OR "DB21".Static_59) AND NOT "DB86".Static_116 AND NOT "DB86".Static_117,
                           Input_6 := "UNO",
                           Input_7 := "DB21".Static_32,
                           Input_8 := "DB21".Static_0,
                           Output_0 => "MV030",
                           Output_2 => "DB32".Static_60,
                           Output_3 => "DB32".Static_61);
END_REGION

REGION Network 8
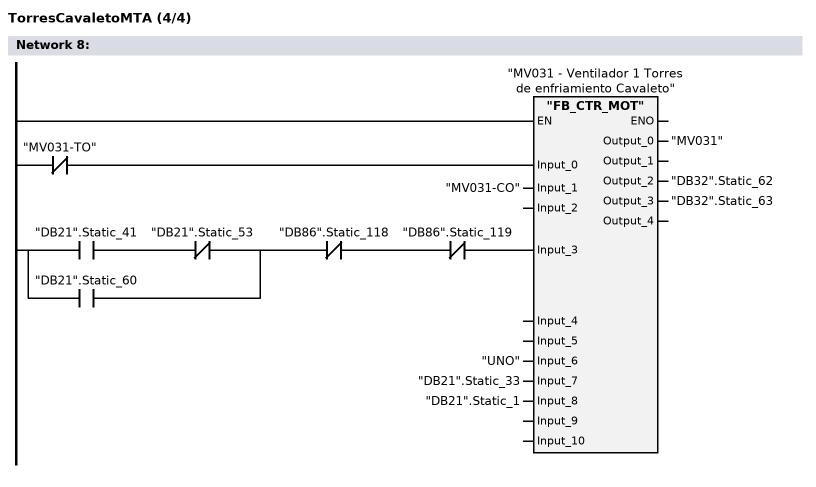
   "MV031 - Ventilador 1 Torres de enfriamiento Cavaleto"(Input_0 := NOT "MV031-TO",   // "FB_CTR_MOT"
                           Input_1 := "MV031-CO",
                           Input_3 := (("DB21".Static_41 AND NOT "DB21".Static_53) OR "DB21".Static_60) AND NOT "DB86".Static_118 AND NOT "DB86".Static_119,
                           Input_6 := "UNO",
                           Input_7 := "DB21".Static_33,
                           Input_8 := "DB21".Static_1,
                           Output_0 => "MV031",
                           Output_2 => "DB32".Static_62,
                           Output_3 => "DB32".Static_63);
END_REGION
END_FUNCTION

// folder: Torres de Agua/Chillers

FUNCTION "TorresAutoMTA" : Void   // FC9, LAD
{ S7_Optimized_Access := 'FALSE' }
VERSION : 0.1
BEGIN

REGION Network 1
